// TIA Portal project "Mes_Con" (V17)

(* hardware
DEVICE "S7-1500/ET200MP station_1"  S7-1500 station
   slot 0: "Rail_0"  Rack  6ES7 590-1***0-0AA0
   slot 1: "PLC_1"  CPU 1515-2 PN  6ES7 515-2AM02-0AB0  V2.9
      slot 3: "CPU display_1"  6ES7591-1BA00-0AA0
      slot 32768: "PROFINET interface_1"  X1
         slot 32769: "Port_1"  X1 P1
         slot 32770: "Port_2"  X1 P2
      slot 33024: "PROFINET interface_2"  X2
         slot 33025: "Port_1"  X2 P1
      slot 34817: "Virtual CP interface port_1"  Virtual CP interface port  Virtual CP interface port
DEVICE "HMI_1"  KTP900 Basic PN
   slot 0: "HMI_1"  KTP900 Basic PN  6AV2 123-2JB03-0AX0  17.0.0.0
   slot 1: "HMI_RT_1"  KTP900 Basic PN  6AV2 123-2JB03-0AX0  17.0.0.0
   slot 5: "HMI_1.IE_CP_1"  PROFINET Interface  17.0.0.0
      slot 1: "PROFINET Interface_1"  PROFINET Interface
         slot 1: "Port_1"  Port
*)

// ===== PLC "PLC_1"  CPU 1515-2 PN =====

VAR_GLOBAL   // PLC tag table "Default tag table"
   "Clock_Byte" AT %MB0 : Byte;
   "Clock_10Hz" AT %M0.0 : Bool;
   "Clock_5Hz" AT %M0.1 : Bool;
   "Clock_2.5Hz" AT %M0.2 : Bool;
   "Clock_2Hz" AT %M0.3 : Bool;
   "Clock_1.25Hz" AT %M0.4 : Bool;
   "Clock_1Hz" AT %M0.5 : Bool;
   "Clock_0.625Hz" AT %M0.6 : Bool;
   "Clock_0.5Hz" AT %M0.7 : Bool;
   "System_Byte" AT %MB1 : Byte;
   "FirstScan" AT %M1.0 : Bool;
   "DiagStatusUpdate" AT %M1.1 : Bool;
   "AlwaysTRUE" AT %M1.2 : Bool;
   "AlwaysFALSE" AT %M1.3 : Bool;
   "PUMP-1_Running" AT %I10.0 : Bool;
   "PUMP-1_Thermic" AT %I10.1 : Bool;
   "PUMP-1_Loc" AT %I10.2 : Bool;
   "PUMP-2_Running" AT %I10.3 : Bool;
   "PUMP-2_Thermic" AT %I10.4 : Bool;
   "PUMP-2_Loc" AT %I10.5 : Bool;
   "PUMP-3_Running" AT %I10.6 : Bool;
   "PUMP-3_Thermic" AT %I10.7 : Bool;
   "PUMP-3_Loc" AT %I11.0 : Bool;
   "PUMP-4_Running" AT %I11.1 : Bool;
   "PUMP-4_Thermic" AT %I11.2 : Bool;
   "PUMP-4_Loc" AT %I11.3 : Bool;
   "Valve-1_Opened" AT %I11.4 : Bool;
   "Valve-1_Closed" AT %I11.5 : Bool;
   "Valve-2_Opened" AT %I11.6 : Bool;
   "Valve-2_Closed" AT %I11.7 : Bool;
   "Valve-3_Opened" AT %I12.0 : Bool;
   "Valve-3_Closed" AT %I12.1 : Bool;
   "Valve-4_Opened" AT %I12.2 : Bool;
   "Valve-4_Closed" AT %I12.3 : Bool;
   "CValve-1_Fbk" AT %IW100 : Word;
   "CValve-2_Fbk" AT %IW102 : Word;
   "CValve-3_Fbk" AT %IW104 : Word;
   "CValve-4_Fbk" AT %IW106 : Word;
   "Pump-1_RPM" AT %IW108 : Word;
   "Pump-2_RPM" AT %IW110 : Word;
   "Pump-3_RPM" AT %IW112 : Word;
   "Pump-4_RPM" AT %IW114 : Word;
   "TT-0001" AT %IW116 : Word;
   "TT-0002" AT %IW118 : Word;
   "PT-0001" AT %IW120 : Word;
   "PT-0002" AT %IW122 : Word;
   "CValve-1_Set" AT %QW200 : Word;
   "CValve-2_Set" AT %QW202 : Word;
   "CValve-3_Set" AT %QW204 : Word;
   "CValve-4_Set" AT %QW206 : Word;
   "Pump-1_SpeedRef" AT %QW208 : Word;
   "Pump-2_SpeedRef" AT %QW210 : Word;
   "Pump-3_SpeedRef" AT %QW212 : Word;
   "Pump-4_SpeedRef" AT %QW214 : Word;
   "Pump-1_Run" AT %Q50.0 : Bool;
   "Pump-2_Run" AT %Q50.1 : Bool;
   "Pump-3_Run" AT %Q50.2 : Bool;
   "Pump-4_Run" AT %Q50.3 : Bool;
   "Valve-1_Open" AT %Q50.4 : Bool;
   "Valve-2_Open" AT %Q50.5 : Bool;
   "Valve-3_Open" AT %Q50.6 : Bool;
   "Valve-4_Open" AT %Q50.7 : Bool;
   "Pump-1_Temp" AT %IW124 : Word;
   "Pump-1_A" AT %IW126 : Word;
   "Pump-2_Temp" AT %IW128 : Word;
   "Pump-2_A" AT %IW130 : Word;
   "Pump-3_Temp" AT %IW132 : Word;
   "Pump-3_A" AT %IW134 : Word;
   "Pump-4_Temp" AT %IW136 : Word;
   "Pump-4_A" AT %IW138 : Word;
END_VAR

TYPE "Popup"
VERSION : 0.1
   STRUCT
      POPUP : Array[0..99] of Bool;
   END_STRUCT;
END_TYPE

TYPE "Valve"
VERSION : 0.1
   STRUCT
      "Mod" : Bool;   // Valf Calisma durumu 0 manuel 1 otomatik
      ManuelOpen : Bool;   // MANUEL START
      ManuelClose : Bool;   // MANUEL STOP
      AutoOpen : Bool;   // AUTO START
      AutoClose : Bool;   // AUTO STOP
      Vana_Open : Bool;   // VANA AÇ
      Vana_Close : Bool;   // VANA KAPAT
      Vana_Opened : Bool;   // VANA AÇIK
      Vana_Closed : Bool;   // VANA KAPALI
      ValveStatus : Int;
      ModStatus : Int;   // VANA STATUS
      ValveIzın : Bool;
      Alarm_Not_Opened : Bool;   // AÇILMIYOR ALRM
      Alarm_Not_Closed : Bool;   // KAPANMIYOR ALARM
      Alarm_Not_Signal : Bool;   // SİNYAL YOK ALARM
      Alarm_Two_Signal : Bool;
      TimeOut : Int;   // ALARM ÇIKIŞ ZAMANI
      Alarm : Bool;   // ALARM
      Alarm_Reset : Bool;   // ALALRM RESET
      PopupClose : Bool;
      PopupInp : Bool;
      Yedek : Bool;
      Yedek_1 : Bool;
      Yedek_2 : Bool;
      Yedek_3 : Bool;
      Yedek_4 : Bool;
      Yedek_5 : Bool;
      Yedek_6 : Bool;
      Yedek_7 : Bool;
      Yedek_8 : Bool;
      Yedek_9 : Bool;
      Yedek_10 : Bool;
      Timer_1 : Int;
      Timer_2 : Int;
      Timer_4 : Int;
      Timer_5 : Int;
      Timer_3 : Int;
      Timer_6 : Int;
      Timer_7 : Int;
      Timer_8 : Int;
      Timer_9 : Int;
   END_STRUCT;
END_TYPE

TYPE "AnalogInput"
VERSION : 0.1
   STRUCT
      Input_Value : Int;
      Input_Value_Conv : Real;
      Mid_Value : Real;
      Measurement_Range : Real;
      "Procces Value_1" : Real;
      Range_Son : Real;
      Measurement_Value_Max : Real;
      Measurement_Value_Min : Real;
      Yedek_2 : Bool;
      Yedek_1 : Bool;
      Range_Control : Bool;
      AlarmTiemOut : Int := 8;
      Timer_1 : Int := 0;
      Timer_2 : Int;
      Alarm : Bool;
      Alarm_Reset : Bool;
      Range_Error : Bool;
   END_STRUCT;
END_TYPE

TYPE "AnalogOutput"
VERSION : 0.1
   STRUCT
      Process_Value : Real;
      Process_Value_Conv : Real;
      Procces_Value_Conv_Int : Int;
      Mid_Valuer : Real;
      Input_Value : Real;
      Input_Value_Real : Real;
      Measurement_Range : Real;
      Measurement_Range_Max : Real;
      Measurement_Range_Min : Real;
      RangeControl : Bool;
      Alarm : Bool;
      Range_Alarm : Bool;
      Alarm_2 : Bool;
      AlarmTimeOut : Int;
      AlarmReset : Bool;
      Yedek : Bool;
      Yedek_1 : Bool;
      Yedek_2 : Bool;
      Yedek_3 : Bool;
      Timer_1 : Int;
      Timer_3 : Int;
      Timer_2 : Int;
   END_STRUCT;
END_TYPE

TYPE "Motor"
VERSION : 0.1
   STRUCT
      "Mod" : Bool;   // 0 = Manuel Mod , 1 = Otomatik Mod
      ManuelStart : Bool;   // HMI Motor Start Button
      ManuelStop : Bool;   // HMI Motor Stop Button
      AutoStart : Bool;   // Logic Auto Start Command
      AutoStop : Bool;   // Logic Auto Stop Command
      "Local/Remote" : Bool;   // Local or Remote Button
      Motor_Rpm : Bool;
      Ucgen_Run : Bool;
      Yildiz_Run : Bool;
      iRunning : Bool;   // Motor Running Information
      iThermic : Bool;   // Motor Thermic Information
      Motor_Izın : Bool;
      Fault : Bool;   // General Fault Information
      Reset : Bool;   // Error Reset Button
      MotorStatus : Int;   // 0=Motor Calismiyor ve Hata Yok 1 = Motor Calisiyor 2 = Motor Calismasini Engelleyen Durum 3 = Motor Arıza Var
      TimeOutAlarm : Bool;   // Motor Timeout Alarm
      ThermicAlarm : Bool;   // Motor Thermic Alarm
      ShortCircuitAlarm : Bool;   // Motor Short Circuit Alarm
      MissingPhaseAlarm : Bool;   // Motor Missing Phase Alarm
      Alarm_Genel : Bool;
      Alarm6 : Bool;
      Alarm7 : Bool;
      Alarm8 : Bool;
      Yedek1 : Bool;
      Yedek2 : Bool;
      Yedek3 : Bool;
      Yedek4 : Bool;
      Yedek5 : Bool;
      Yedek6 : Bool;
      Yedek7 : Bool;
      Timer1 : Int;
      Timer2 : Int;
      Timer3 : Int;
      Timer4 : Int;
      Timer5 : Int;
      Timer6 : Int;
   END_STRUCT;
END_TYPE

TYPE "ElValve"
VERSION : 0.1
   STRUCT
      VanaOpened : Bool;
      VanaClosed : Bool;
      VanaAlarm : Bool;
      Alarm_Not_Signal : Bool;   // SİNYAL YOK ALARM
      Alarm_Two_Signal : Bool;
      Alarm_Genel : Bool;
      Alarm_Reset : Bool;
      ElV_Status : Int;
      Yedek_1 : Bool;
      Yedek_2 : Bool;
      Yedek_3 : Bool;
      Timer_1 : Int;
      Timer_2 : Int;
      Timer_3 : Int;
      TimeOut : Int;
   END_STRUCT;
END_TYPE

TYPE "FM"
VERSION : 0.1
   STRUCT
      P_Value : Real;
      Flow_Pulse_N : Int;
      F_Pulse : Bool;
      Pulse_Kg : Real;
      Total_Value : DInt;
      Set_Value : DInt;
      Tank_Value : DInt;
      TankBosaltıldı : Bool;
      SU_Alım_Run : Bool;
      TankValue_Reset : Bool;
      Total_Value_Reset : Bool;
      Pulse_Reset : Bool;
      Yedek : Bool;
      Yedek_1 : Bool;
      Yedek_2 : Int;
      Yedek_3 : Int;
   END_STRUCT;
END_TYPE

TYPE "Gunler"
VERSION : 0.1
   STRUCT
      Pazartesi : Bool;
      Salı : Bool;
      Çarşamba : Bool;
      Perşembe : Bool;
      Cuma : Bool;
      Cumartesi : Bool;
      Pazar : Bool;
      Pazartesi_Veri : Int;
      Salı_Veri : Int;
      Çarşamba_Veri : Int;
      Perşembe_Veri : Int;
      Cuma_Veri : Int;
      Cumartesi_Veri : Int;
      Pazar_Veri : Int;
      Yedek : Bool;
      Yedek_1 : Bool;
      Yedek_2 : Bool;
      Yedek_3 : Bool;
      Yedek_4 : Bool;
      Yedek_5 : Bool;
      Yedek_6 : Bool;
      Yedek_7 : Bool;
      "Timer" : Int;
      Timer_1 : Int;
      Timer_2 : Int;
      Timer_3 : Int;
   END_STRUCT;
END_TYPE

// folder: Data

DATA_BLOCK "Sim"   // DB5
{ S7_Optimized_Access := 'TRUE' }
VERSION : 0.1
   VAR
      "SPUMP-1_Running" : Bool;
      "SPUMP-1_Thermic" : Bool;
      "SPUMP-1_Loc" : Bool;
      "SPUMP-2_Running" : Bool;
      "SPUMP-2_Thermic" : Bool;
      "SPUMP-2_Loc" : Bool;
      "SPUMP-3_Running" : Bool;
      "SPUMP-3_Thermic" : Bool;
      "SPUMP-3_Loc" : Bool;
      "SPUMP-4_Running" : Bool;
      "SPUMP-4_Thermic" : Bool;
      "SPUMP-4_Loc" : Bool;
      "SValve-1_Opened" : Bool;
      "SValve-1_Closed" : Bool;
      "SValve-2_Opened" : Bool;
      "SValve-2_Closed" : Bool;
      "SValve-3_Opened" : Bool;
      "SValve-3_Closed" : Bool;
      "SValve-4_Opened" : Bool;
      "SValve-4_Closed" : Bool;
      "SPump-1_Run" : Bool;
      "SPump-2_Run" : Bool;
      "SPump-3_Run" : Bool;
      "SPump-4_Run" : Bool;
      "SValve-1_Open" : Bool;
      "SValve-2_Open" : Bool;
      "SValve-3_Open" : Bool;
      "SValve-4_Open" : Bool;
      "SCValve-1_Fbk" : Word;
      "SCValve-2_Fbk" : Word;
      "SCValve-3_Fbk" : Word;
      "SCValve-4_Fbk" : Word;
      "SPump-1_RPM" : Word;
      "SPump-2_RPM" : Word;
      "SPump-3_RPM" : Word;
      "SPump-4_RPM" : Word;
      "SPump-1_Temp" : Word;
      "SPump-1_A" : Word;
      "SPump-2_Temp" : Word;
      "SPump-2_A" : Word;
      "SPump-3_Temp" : Word;
      "SPump-3_A" : Word;
      "SPump-4_Temp" : Word;
      "SPump-4_A" : Word;
      "STT-0001" : Word;
      "STT-0002" : Word;
      "SPT-0001" : Word;
      "SPT-0002" : Word;
      "SCValve-1_Set" : Word;
      "SCValve-2_Set" : Word;
      "SCValve-3_Set" : Word;
      "SCValve-4_Set" : Word;
      "SPump-1_SpeedRef" : Word;
      "SPump-2_SpeedRef" : Word;
      "SPump-3_SpeedRef" : Word;
      "SPump-4_SpeedRef" : Word;
      SİM_MOD : Bool;
   END_VAR
BEGIN
END_DATA_BLOCK

// folder: Data/Eqp

DATA_BLOCK "PUMP"   // DB1
{ S7_Optimized_Access := 'TRUE' }
VERSION : 0.1
   VAR
      "PUMP-1" : "Motor";
      "PUMP-2" : "Motor";
      "PUMP-3" : "Motor";
      "PUMP-4" : "Motor";
   END_VAR
BEGIN
END_DATA_BLOCK

DATA_BLOCK "VALVE-H"   // DB2
{ S7_Optimized_Access := 'TRUE' }
VERSION : 0.1
   VAR
      "VALVE-1" : "Valve";
      "VALVE-2" : "Valve";
      "VALVE-3" : "Valve";
      "VALVE-4" : "Valve";
   END_VAR
BEGIN
END_DATA_BLOCK

DATA_BLOCK "VALVE-C"   // DB3
{ S7_Optimized_Access := 'TRUE' }
VERSION : 0.1
   VAR
      "CONTROLV-1" : "AnalogOutput";
      "CONTROLV-2" : "AnalogOutput";
      "CONTROLV-3" : "AnalogOutput";
      "CONTROLV-4" : "AnalogOutput";
   END_VAR
BEGIN
END_DATA_BLOCK

DATA_BLOCK "TT-PT"   // DB4
{ S7_Optimized_Access := 'TRUE' }
VERSION : 0.1
   VAR
      "TT-0001" : "AnalogInput";
      "TT-0002" : "AnalogInput";
      "PT-0001" : "AnalogInput";
      "PT-0002" : "AnalogInput";
   END_VAR
BEGIN
END_DATA_BLOCK

// folder: Data/HMI

DATA_BLOCK "HMI"   // DB7
{ S7_Optimized_Access := 'TRUE' }
VERSION : 0.1
   VAR
      Popup : "Popup";
      "CValve-1_Set" : Int;
      "CValve-2_Set" : Int;
      "CValve-3_Set" : Int;
      "CValve-4_Set" : Int;
      "Pump-1" : Int;
      "Pump-2" : Int;
      "Pump-3" : Int;
      "Pump-4" : Int;
   END_VAR
BEGIN
END_DATA_BLOCK

// folder: Data/mes

DATA_BLOCK "Connection"   // DB6
{ S7_Optimized_Access := 'FALSE' }
VERSION : 0.1
   VAR
      "CV-1Flt" : Bool;
      "CV-2Flt" : Bool;
      "CV-3Flt" : Bool;
      "CV-4Flt" : Bool;
      "TT1-FLT" : Bool;
      "TT2-FLT" : Bool;
      "PT1-FLT" : Bool;
      "PT2-FLT" : Bool;
      "Pump-1Status" : Word;
      "Pump-2Status" : Word;
      "Pump-3Status" : Word;
      "Pump-4Status" : Word;
      "V1-Status" : Word;
      "V2-Status" : Word;
      "V3-Status" : Word;
      "V4-Status" : Word;
      "Pump1-Rpm" : Word;
      "Pump2-Rpm" : Word;
      "Pump3-Rpm" : Word;
      "Pump4-Rpm" : Word;
      "CV1-Percent" : Word;
      "CV2-Percent" : Word;
      "CV3-Percent" : Word;
      "CV4-Percent" : Word;
      "TT1-Value" : Word;
      "TT2-Value" : Word;
      "PT1-Value" : Word;
      "PT2-Value" : Word;
   END_VAR
BEGIN
END_DATA_BLOCK

DATA_BLOCK "workorder"   // DB10
{ S7_Optimized_Access := 'FALSE' }
VERSION : 0.1
   VAR
      "Work_Order-1_Active" : Bool;
      "Work_Order-2_Active" : Bool;
      "Work_Order-3_Active" : Bool;
      "Work_Order-4_Active" : Bool;
      "Work_Order-5_Active" : Bool;
      "Work_Order-6_Active" : Bool;
      "Work_Order-7_Active" : Bool;
      "Work_Order-8_Active" : Bool;
      "Work_Order-9_Active" : Bool;
      "Work_Order-10_Active" : Bool;
      "Work_Order-11_Active" : Bool;
      "Work_Order-12_Active" : Bool;
      "Work_Order-13_Active" : Bool;
      "Work_Order-14_Active" : Bool;
      "Work_Order-15_Active" : Bool;
   END_VAR
BEGIN
END_DATA_BLOCK

DATA_BLOCK "maint"   // DB100
{ S7_Optimized_Access := 'TRUE' }
VERSION : 0.1
   VAR
      "Pump-1_Sim" : Bool;
      "Pump-1_Running" : Bool;
      "Pump-1_Loc" : Bool;
      "Pump-1_PhaseAlarm" : Bool;
      "Pump-1_ThermicAlarm" : Bool;
      "Pump-1_TimeOutAlarm" : Bool;
      "Pump-1_ShortCircuit" : Bool;
      "Pump-2_Sim" : Bool;
      "Pump-2_Running" : Bool;
      "Pump-2_Loc" : Bool;
      "Pump-2_PhaseAlarm" : Bool;
      "Pump-2_ThermicAlarm" : Bool;
      "Pump-2_TimeOutAlarm" : Bool;
      "Pump-2_ShortCircuit" : Bool;
      "Pump-3_Sim" : Bool;
      "Pump-3_Running" : Bool;
      "Pump-3_Loc" : Bool;
      "Pump-3_PhaseAlarm" : Bool;
      "Pump-3_ThermicAlarm" : Bool;
      "Pump-3_TimeOutAlarm" : Bool;
      "Pump-3_ShortCircuit" : Bool;
      "Pump-4_Sim" : Bool;
      "Pump-4_Running" : Bool;
      "Pump-4_Loc" : Bool;
      "Pump-4_PhaseAlarm" : Bool;
      "Pump-4_ThermicAlarm" : Bool;
      "Pump-4_TimeOutAlarm" : Bool;
      "Pump-4_ShortCircuit" : Bool;
      "Valve-1_Sim" : Bool;
      "Valve-1_NotOpened" : Bool;
      "Valve-1_NotClosed" : Bool;
      "Valve-1_NotSignal" : Bool;
      "Valve-1_TwoSignal" : Bool;
      "Valve-2_Sim" : Bool;
      "Valve-2_NotOpened" : Bool;
      "Valve-2_NotClosed" : Bool;
      "Valve-2_NotSignal" : Bool;
      "Valve-2_TwoSignal" : Bool;
      "Valve-3_Sim" : Bool;
      "Valve-3_NotOpened" : Bool;
      "Valve-3_NotClosed" : Bool;
      "Valve-3_NotSignal" : Bool;
      "Valve-3_TwoSignal" : Bool;
      "Valve-4_Sim" : Bool;
      "Valve-4_NotOpened" : Bool;
      "Valve-4_NotClosed" : Bool;
      "Valve-4_NotSignal" : Bool;
      "Valve-4_TwoSignal" : Bool;
      "Pump-1_A" : Word;
      "Pump-1_Temp" : Word;
      "Pump-2_A" : Word;
      "Pump-2_Temp" : Word;
      "Pump-3_A" : Word;
      "Pump-3_Temp" : Word;
      "Pump-4_A" : Word;
      "Pump-4_Temp" : Word;
      "TT-0001" : Word;
      "TT-0002" : Word;
      "PT-0001" : Word;
      "PT-0002" : Word;
      "CValve-1_FBK" : Word;
      "CValve-2_FBK" : Word;
      "CValve-3_FBK" : Word;
      "CValve-4_FBK" : Word;
   END_VAR
BEGIN
END_DATA_BLOCK

// folder: (top level)

FUNCTION "Equipment" : Void   // FC2, LAD
{ S7_Optimized_Access := 'TRUE' }
VERSION : 0.1
BEGIN

REGION Network 1: PUMP-1
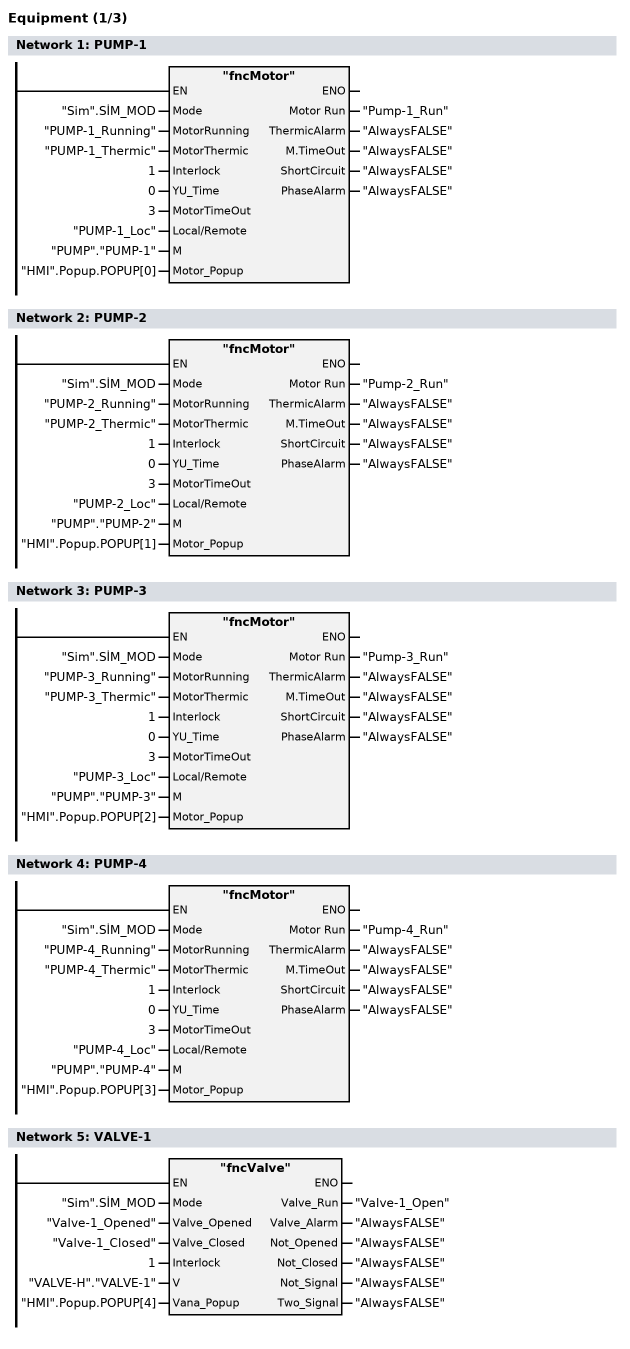
   RUNG wire#powerrail
      "fncMotor"(Mode := "Sim".SİM_MOD, MotorRunning := "PUMP-1_Running", MotorThermic := "PUMP-1_Thermic", Interlock := 1, YU_Time := 0, MotorTimeOut := 3, "Local/Remote" := "PUMP-1_Loc", "M" := "PUMP"."PUMP-1", Motor_Popup := "HMI".Popup.POPUP[0], "Motor Run" => "Pump-1_Run", ThermicAlarm => "AlwaysFALSE", "M.TimeOut" => "AlwaysFALSE", ShortCircuit => "AlwaysFALSE", PhaseAlarm => "AlwaysFALSE")
   END_RUNG
   // the same network as SCL:
   "fncMotor"(Mode := "Sim".SİM_MOD,
              MotorRunning := "PUMP-1_Running",
              MotorThermic := "PUMP-1_Thermic",
              Interlock := 1,
              YU_Time := 0,
              MotorTimeOut := 3,
              "Local/Remote" := "PUMP-1_Loc",
              "M" := "PUMP"."PUMP-1",
              Motor_Popup := "HMI".Popup.POPUP[0],
              "Motor Run" => "Pump-1_Run",
              ThermicAlarm => "AlwaysFALSE",
              "M.TimeOut" => "AlwaysFALSE",
              ShortCircuit => "AlwaysFALSE",
              PhaseAlarm => "AlwaysFALSE");
END_REGION

REGION Network 2: PUMP-2
   RUNG wire#powerrail
      "fncMotor"(Mode := "Sim".SİM_MOD, MotorRunning := "PUMP-2_Running", MotorThermic := "PUMP-2_Thermic", Interlock := 1, YU_Time := 0, MotorTimeOut := 3, "Local/Remote" := "PUMP-2_Loc", "M" := "PUMP"."PUMP-2", Motor_Popup := "HMI".Popup.POPUP[1], "Motor Run" => "Pump-2_Run", ThermicAlarm => "AlwaysFALSE", "M.TimeOut" => "AlwaysFALSE", ShortCircuit => "AlwaysFALSE", PhaseAlarm => "AlwaysFALSE")
   END_RUNG
   // the same network as SCL:
   "fncMotor"(Mode := "Sim".SİM_MOD,
              MotorRunning := "PUMP-2_Running",
              MotorThermic := "PUMP-2_Thermic",
              Interlock := 1,
              YU_Time := 0,
              MotorTimeOut := 3,
              "Local/Remote" := "PUMP-2_Loc",
              "M" := "PUMP"."PUMP-2",
              Motor_Popup := "HMI".Popup.POPUP[1],
              "Motor Run" => "Pump-2_Run",
              ThermicAlarm => "AlwaysFALSE",
              "M.TimeOut" => "AlwaysFALSE",
              ShortCircuit => "AlwaysFALSE",
              PhaseAlarm => "AlwaysFALSE");
END_REGION

REGION Network 3: PUMP-3
   RUNG wire#powerrail
      "fncMotor"(Mode := "Sim".SİM_MOD, MotorRunning := "PUMP-3_Running", MotorThermic := "PUMP-3_Thermic", Interlock := 1, YU_Time := 0, MotorTimeOut := 3, "Local/Remote" := "PUMP-3_Loc", "M" := "PUMP"."PUMP-3", Motor_Popup := "HMI".Popup.POPUP[2], "Motor Run" => "Pump-3_Run", ThermicAlarm => "AlwaysFALSE", "M.TimeOut" => "AlwaysFALSE", ShortCircuit => "AlwaysFALSE", PhaseAlarm => "AlwaysFALSE")
   END_RUNG
   // the same network as SCL:
   "fncMotor"(Mode := "Sim".SİM_MOD,
              MotorRunning := "PUMP-3_Running",
              MotorThermic := "PUMP-3_Thermic",
              Interlock := 1,
              YU_Time := 0,
              MotorTimeOut := 3,
              "Local/Remote" := "PUMP-3_Loc",
              "M" := "PUMP"."PUMP-3",
              Motor_Popup := "HMI".Popup.POPUP[2],
              "Motor Run" => "Pump-3_Run",
              ThermicAlarm => "AlwaysFALSE",
              "M.TimeOut" => "AlwaysFALSE",
              ShortCircuit => "AlwaysFALSE",
              PhaseAlarm => "AlwaysFALSE");
END_REGION

REGION Network 4: PUMP-4
   RUNG wire#powerrail
      "fncMotor"(Mode := "Sim".SİM_MOD, MotorRunning := "PUMP-4_Running", MotorThermic := "PUMP-4_Thermic", Interlock := 1, YU_Time := 0, MotorTimeOut := 3, "Local/Remote" := "PUMP-4_Loc", "M" := "PUMP"."PUMP-4", Motor_Popup := "HMI".Popup.POPUP[3], "Motor Run" => "Pump-4_Run", ThermicAlarm => "AlwaysFALSE", "M.TimeOut" => "AlwaysFALSE", ShortCircuit => "AlwaysFALSE", PhaseAlarm => "AlwaysFALSE")
   END_RUNG
   // the same network as SCL:
   "fncMotor"(Mode := "Sim".SİM_MOD,
              MotorRunning := "PUMP-4_Running",
              MotorThermic := "PUMP-4_Thermic",
              Interlock := 1,
              YU_Time := 0,
              MotorTimeOut := 3,
              "Local/Remote" := "PUMP-4_Loc",
              "M" := "PUMP"."PUMP-4",
              Motor_Popup := "HMI".Popup.POPUP[3],
              "Motor Run" => "Pump-4_Run",
              ThermicAlarm => "AlwaysFALSE",
              "M.TimeOut" => "AlwaysFALSE",
              ShortCircuit => "AlwaysFALSE",
              PhaseAlarm => "AlwaysFALSE");
END_REGION

REGION Network 5: VALVE-1
   RUNG wire#powerrail
      "fncValve"(Mode := "Sim".SİM_MOD, Valve_Opened := "Valve-1_Opened", Valve_Closed := "Valve-1_Closed", Interlock := 1, V := "VALVE-H"."VALVE-1", Vana_Popup := "HMI".Popup.POPUP[4], Valve_Run => "Valve-1_Open", Valve_Alarm => "AlwaysFALSE", Not_Opened => "AlwaysFALSE", Not_Closed => "AlwaysFALSE", Not_Signal => "AlwaysFALSE", Two_Signal => "AlwaysFALSE")
   END_RUNG
   // the same network as SCL:
   "fncValve"(Mode := "Sim".SİM_MOD,
              Valve_Opened := "Valve-1_Opened",
              Valve_Closed := "Valve-1_Closed",
              Interlock := 1,
              V := "VALVE-H"."VALVE-1",
              Vana_Popup := "HMI".Popup.POPUP[4],
              Valve_Run => "Valve-1_Open",
              Valve_Alarm => "AlwaysFALSE",
              Not_Opened => "AlwaysFALSE",
              Not_Closed => "AlwaysFALSE",
              Not_Signal => "AlwaysFALSE",
              Two_Signal => "AlwaysFALSE");
END_REGION

REGION Network 6: VALVE-2
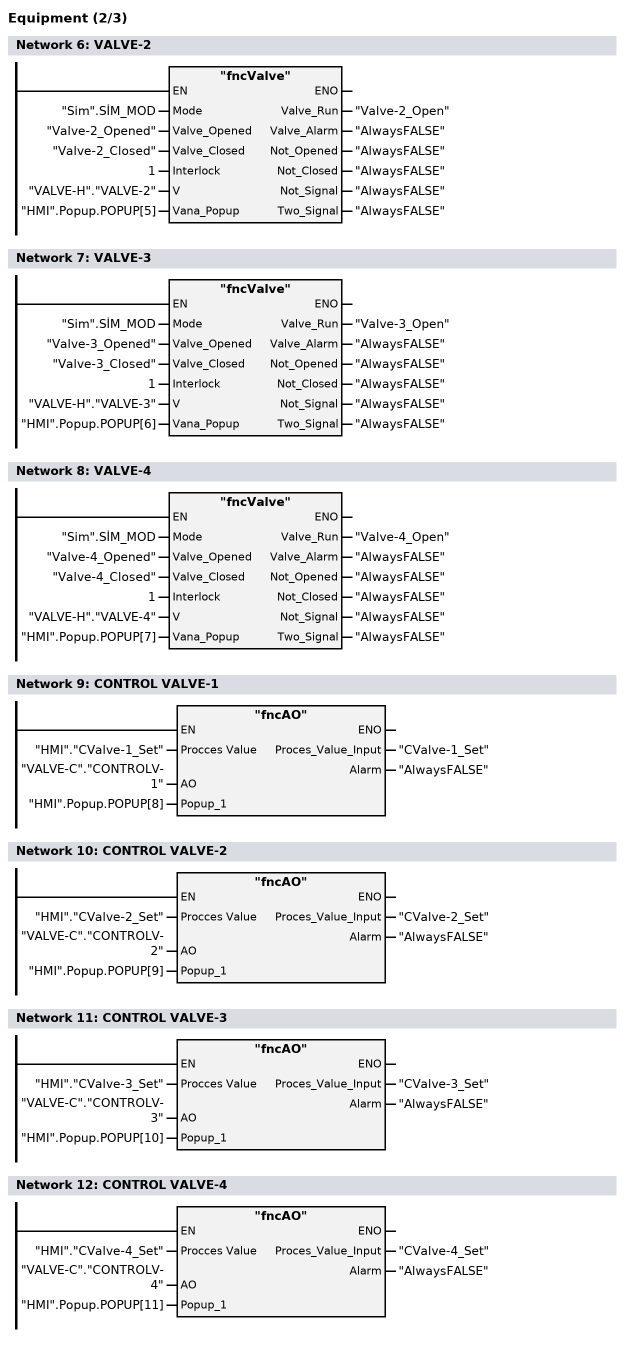
   RUNG wire#powerrail
      "fncValve"(Mode := "Sim".SİM_MOD, Valve_Opened := "Valve-2_Opened", Valve_Closed := "Valve-2_Closed", Interlock := 1, V := "VALVE-H"."VALVE-2", Vana_Popup := "HMI".Popup.POPUP[5], Valve_Run => "Valve-2_Open", Valve_Alarm => "AlwaysFALSE", Not_Opened => "AlwaysFALSE", Not_Closed => "AlwaysFALSE", Not_Signal => "AlwaysFALSE", Two_Signal => "AlwaysFALSE")
   END_RUNG
   // the same network as SCL:
   "fncValve"(Mode := "Sim".SİM_MOD,
              Valve_Opened := "Valve-2_Opened",
              Valve_Closed := "Valve-2_Closed",
              Interlock := 1,
              V := "VALVE-H"."VALVE-2",
              Vana_Popup := "HMI".Popup.POPUP[5],
              Valve_Run => "Valve-2_Open",
              Valve_Alarm => "AlwaysFALSE",
              Not_Opened => "AlwaysFALSE",
              Not_Closed => "AlwaysFALSE",
              Not_Signal => "AlwaysFALSE",
              Two_Signal => "AlwaysFALSE");
END_REGION

REGION Network 7: VALVE-3
   RUNG wire#powerrail
      "fncValve"(Mode := "Sim".SİM_MOD, Valve_Opened := "Valve-3_Opened", Valve_Closed := "Valve-3_Closed", Interlock := 1, V := "VALVE-H"."VALVE-3", Vana_Popup := "HMI".Popup.POPUP[6], Valve_Run => "Valve-3_Open", Valve_Alarm => "AlwaysFALSE", Not_Opened => "AlwaysFALSE", Not_Closed => "AlwaysFALSE", Not_Signal => "AlwaysFALSE", Two_Signal => "AlwaysFALSE")
   END_RUNG
   // the same network as SCL:
   "fncValve"(Mode := "Sim".SİM_MOD,
              Valve_Opened := "Valve-3_Opened",
              Valve_Closed := "Valve-3_Closed",
              Interlock := 1,
              V := "VALVE-H"."VALVE-3",
              Vana_Popup := "HMI".Popup.POPUP[6],
              Valve_Run => "Valve-3_Open",
              Valve_Alarm => "AlwaysFALSE",
              Not_Opened => "AlwaysFALSE",
              Not_Closed => "AlwaysFALSE",
              Not_Signal => "AlwaysFALSE",
              Two_Signal => "AlwaysFALSE");
END_REGION

REGION Network 8: VALVE-4
   RUNG wire#powerrail
      "fncValve"(Mode := "Sim".SİM_MOD, Valve_Opened := "Valve-4_Opened", Valve_Closed := "Valve-4_Closed", Interlock := 1, V := "VALVE-H"."VALVE-4", Vana_Popup := "HMI".Popup.POPUP[7], Valve_Run => "Valve-4_Open", Valve_Alarm => "AlwaysFALSE", Not_Opened => "AlwaysFALSE", Not_Closed => "AlwaysFALSE", Not_Signal => "AlwaysFALSE", Two_Signal => "AlwaysFALSE")
   END_RUNG
   // the same network as SCL:
   "fncValve"(Mode := "Sim".SİM_MOD,
              Valve_Opened := "Valve-4_Opened",
              Valve_Closed := "Valve-4_Closed",
              Interlock := 1,
              V := "VALVE-H"."VALVE-4",
              Vana_Popup := "HMI".Popup.POPUP[7],
              Valve_Run => "Valve-4_Open",
              Valve_Alarm => "AlwaysFALSE",
              Not_Opened => "AlwaysFALSE",
              Not_Closed => "AlwaysFALSE",
              Not_Signal => "AlwaysFALSE",
              Two_Signal => "AlwaysFALSE");
END_REGION

REGION Network 9: CONTROL VALVE-1
   RUNG wire#powerrail
      "fncAO"("Procces Value" := "HMI"."CValve-1_Set", AO := "VALVE-C"."CONTROLV-1", Popup_1 := "HMI".Popup.POPUP[8], Proces_Value_Input => "CValve-1_Set", Alarm => "AlwaysFALSE")
   END_RUNG
   // the same network as SCL:
   "fncAO"("Procces Value" := "HMI"."CValve-1_Set",
           AO := "VALVE-C"."CONTROLV-1",
           Popup_1 := "HMI".Popup.POPUP[8],
           Proces_Value_Input => "CValve-1_Set",
           Alarm => "AlwaysFALSE");
END_REGION

REGION Network 10: CONTROL VALVE-2
   RUNG wire#powerrail
      "fncAO"("Procces Value" := "HMI"."CValve-2_Set", AO := "VALVE-C"."CONTROLV-2", Popup_1 := "HMI".Popup.POPUP[9], Proces_Value_Input => "CValve-2_Set", Alarm => "AlwaysFALSE")
   END_RUNG
   // the same network as SCL:
   "fncAO"("Procces Value" := "HMI"."CValve-2_Set",
           AO := "VALVE-C"."CONTROLV-2",
           Popup_1 := "HMI".Popup.POPUP[9],
           Proces_Value_Input => "CValve-2_Set",
           Alarm => "AlwaysFALSE");
END_REGION

REGION Network 11: CONTROL VALVE-3
   RUNG wire#powerrail
      "fncAO"("Procces Value" := "HMI"."CValve-3_Set", AO := "VALVE-C"."CONTROLV-3", Popup_1 := "HMI".Popup.POPUP[10], Proces_Value_Input => "CValve-3_Set", Alarm => "AlwaysFALSE")
   END_RUNG
   // the same network as SCL:
   "fncAO"("Procces Value" := "HMI"."CValve-3_Set",
           AO := "VALVE-C"."CONTROLV-3",
           Popup_1 := "HMI".Popup.POPUP[10],
           Proces_Value_Input => "CValve-3_Set",
           Alarm => "AlwaysFALSE");
END_REGION

REGION Network 12: CONTROL VALVE-4
   RUNG wire#powerrail
      "fncAO"("Procces Value" := "HMI"."CValve-4_Set", AO := "VALVE-C"."CONTROLV-4", Popup_1 := "HMI".Popup.POPUP[11], Proces_Value_Input => "CValve-4_Set", Alarm => "AlwaysFALSE")
   END_RUNG
   // the same network as SCL:
   "fncAO"("Procces Value" := "HMI"."CValve-4_Set",
           AO := "VALVE-C"."CONTROLV-4",
           Popup_1 := "HMI".Popup.POPUP[11],
           Proces_Value_Input => "CValve-4_Set",
           Alarm => "AlwaysFALSE");
END_REGION

REGION Network 13: TT-0001
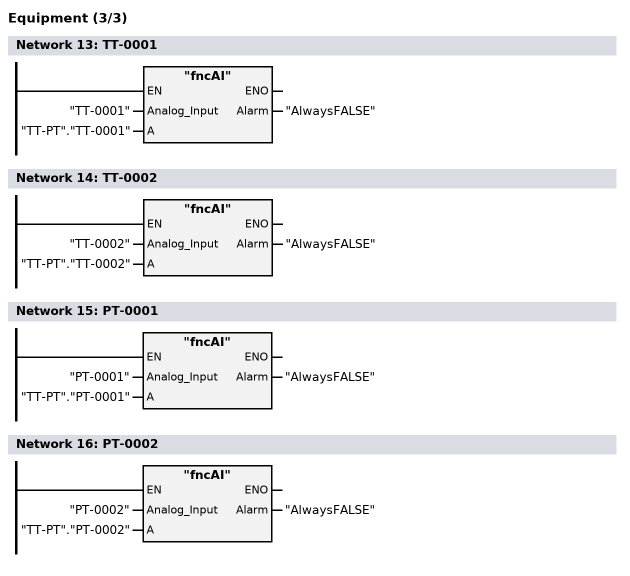
   RUNG wire#powerrail
      "fncAI"(Analog_Input := "TT-0001", "A" := "TT-PT"."TT-0001", Alarm => "AlwaysFALSE")
   END_RUNG
   // the same network as SCL:
   "fncAI"(Analog_Input := "TT-0001", "A" := "TT-PT"."TT-0001", Alarm => "AlwaysFALSE");
END_REGION

REGION Network 14: TT-0002
   RUNG wire#powerrail
      "fncAI"(Analog_Input := "TT-0002", "A" := "TT-PT"."TT-0002", Alarm => "AlwaysFALSE")
   END_RUNG
   // the same network as SCL:
   "fncAI"(Analog_Input := "TT-0002", "A" := "TT-PT"."TT-0002", Alarm => "AlwaysFALSE");
END_REGION

REGION Network 15: PT-0001
   RUNG wire#powerrail
      "fncAI"(Analog_Input := "PT-0001", "A" := "TT-PT"."PT-0001", Alarm => "AlwaysFALSE")
   END_RUNG
   // the same network as SCL:
   "fncAI"(Analog_Input := "PT-0001", "A" := "TT-PT"."PT-0001", Alarm => "AlwaysFALSE");
END_REGION

REGION Network 16: PT-0002
   RUNG wire#powerrail
      "fncAI"(Analog_Input := "PT-0002", "A" := "TT-PT"."PT-0002", Alarm => "AlwaysFALSE")
   END_RUNG
   // the same network as SCL:
   "fncAI"(Analog_Input := "PT-0002", "A" := "TT-PT"."PT-0002", Alarm => "AlwaysFALSE");
END_REGION
END_FUNCTION

FUNCTION "Simfnc" : Void   // FC19, LAD
{ S7_Optimized_Access := 'TRUE' }
VERSION : 0.1
BEGIN

REGION Network 1: PUMP-1
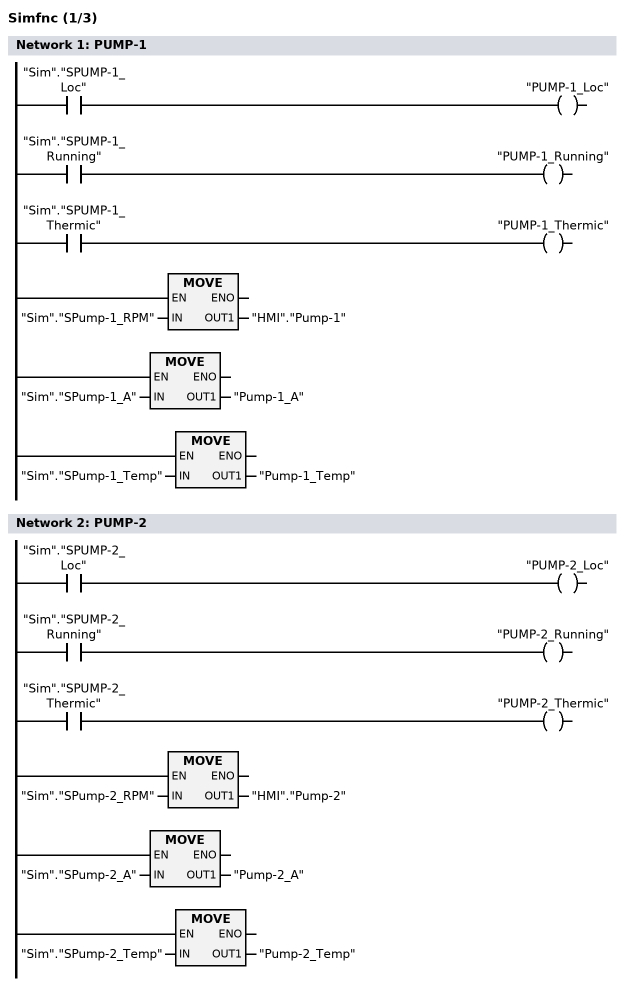
   RUNG wire#powerrail
      Contact( "Sim"."SPUMP-1_Loc" )
      Coil( "PUMP-1_Loc" )
   END_RUNG
   RUNG wire#powerrail
      Contact( "Sim"."SPUMP-1_Running" )
      Coil( "PUMP-1_Running" )
   END_RUNG
   RUNG wire#powerrail
      Contact( "Sim"."SPUMP-1_Thermic" )
      Coil( "PUMP-1_Thermic" )
   END_RUNG
   RUNG wire#powerrail
      Move(in := "Sim"."SPump-1_RPM", out1 => "HMI"."Pump-1")
   END_RUNG
   RUNG wire#powerrail
      Move(in := "Sim"."SPump-1_A", out1 => "Pump-1_A")
   END_RUNG
   RUNG wire#powerrail
      Move(in := "Sim"."SPump-1_Temp", out1 => "Pump-1_Temp")
   END_RUNG
   // the same network as SCL:
   "PUMP-1_Loc" := "Sim"."SPUMP-1_Loc";
   "PUMP-1_Running" := "Sim"."SPUMP-1_Running";
   "PUMP-1_Thermic" := "Sim"."SPUMP-1_Thermic";
   "HMI"."Pump-1" := "Sim"."SPump-1_RPM";
   "Pump-1_A" := "Sim"."SPump-1_A";
   "Pump-1_Temp" := "Sim"."SPump-1_Temp";
END_REGION

REGION Network 2: PUMP-2
   RUNG wire#powerrail
      Contact( "Sim"."SPUMP-2_Loc" )
      Coil( "PUMP-2_Loc" )
   END_RUNG
   RUNG wire#powerrail
      Contact( "Sim"."SPUMP-2_Running" )
      Coil( "PUMP-2_Running" )
   END_RUNG
   RUNG wire#powerrail
      Contact( "Sim"."SPUMP-2_Thermic" )
      Coil( "PUMP-2_Thermic" )
   END_RUNG
   RUNG wire#powerrail
      Move(in := "Sim"."SPump-2_RPM", out1 => "HMI"."Pump-2")
   END_RUNG
   RUNG wire#powerrail
      Move(in := "Sim"."SPump-2_A", out1 => "Pump-2_A")
   END_RUNG
   RUNG wire#powerrail
      Move(in := "Sim"."SPump-2_Temp", out1 => "Pump-2_Temp")
   END_RUNG
   // the same network as SCL:
   "PUMP-2_Loc" := "Sim"."SPUMP-2_Loc";
   "PUMP-2_Running" := "Sim"."SPUMP-2_Running";
   "PUMP-2_Thermic" := "Sim"."SPUMP-2_Thermic";
   "HMI"."Pump-2" := "Sim"."SPump-2_RPM";
   "Pump-2_A" := "Sim"."SPump-2_A";
   "Pump-2_Temp" := "Sim"."SPump-2_Temp";
END_REGION

REGION Network 3: PUMP-3
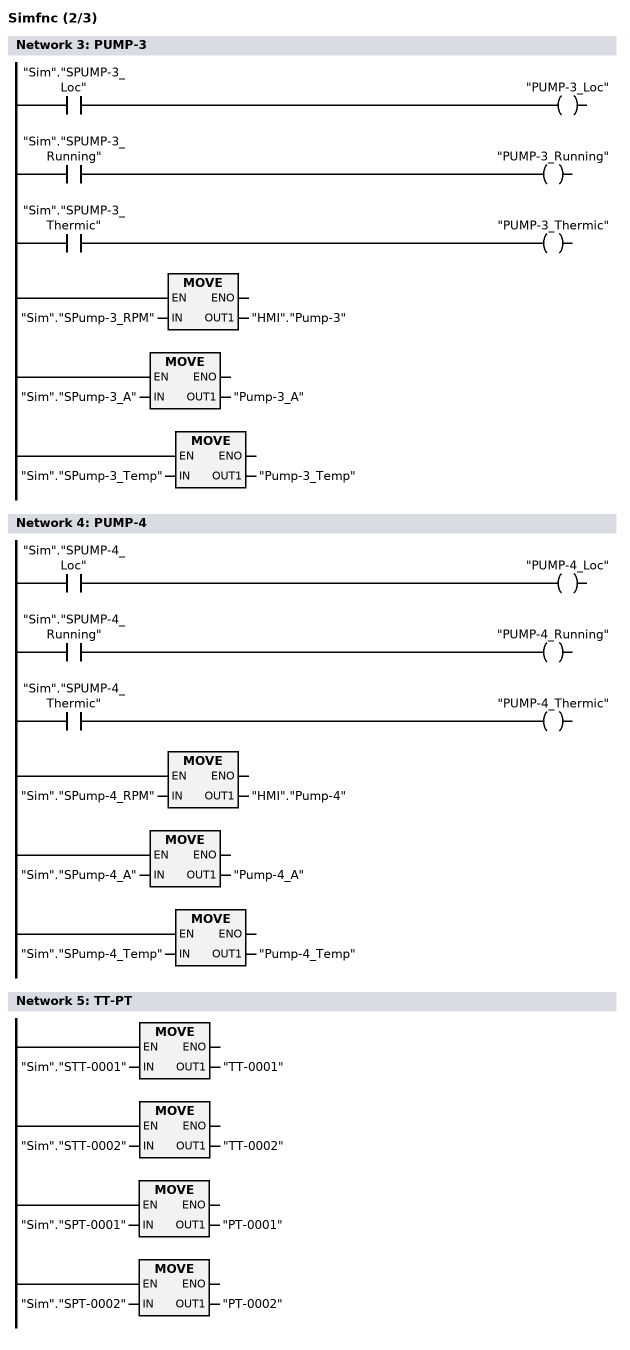
   RUNG wire#powerrail
      Contact( "Sim"."SPUMP-3_Loc" )
      Coil( "PUMP-3_Loc" )
   END_RUNG
   RUNG wire#powerrail
      Contact( "Sim"."SPUMP-3_Running" )
      Coil( "PUMP-3_Running" )
   END_RUNG
   RUNG wire#powerrail
      Contact( "Sim"."SPUMP-3_Thermic" )
      Coil( "PUMP-3_Thermic" )
   END_RUNG
   RUNG wire#powerrail
      Move(in := "Sim"."SPump-3_RPM", out1 => "HMI"."Pump-3")
   END_RUNG
   RUNG wire#powerrail
      Move(in := "Sim"."SPump-3_A", out1 => "Pump-3_A")
   END_RUNG
   RUNG wire#powerrail
      Move(in := "Sim"."SPump-3_Temp", out1 => "Pump-3_Temp")
   END_RUNG
   // the same network as SCL:
   "PUMP-3_Loc" := "Sim"."SPUMP-3_Loc";
   "PUMP-3_Running" := "Sim"."SPUMP-3_Running";
   "PUMP-3_Thermic" := "Sim"."SPUMP-3_Thermic";
   "HMI"."Pump-3" := "Sim"."SPump-3_RPM";
   "Pump-3_A" := "Sim"."SPump-3_A";
   "Pump-3_Temp" := "Sim"."SPump-3_Temp";
END_REGION

REGION Network 4: PUMP-4
   RUNG wire#powerrail
      Contact( "Sim"."SPUMP-4_Loc" )
      Coil( "PUMP-4_Loc" )
   END_RUNG
   RUNG wire#powerrail
      Contact( "Sim"."SPUMP-4_Running" )
      Coil( "PUMP-4_Running" )
   END_RUNG
   RUNG wire#powerrail
      Contact( "Sim"."SPUMP-4_Thermic" )
      Coil( "PUMP-4_Thermic" )
   END_RUNG
   RUNG wire#powerrail
      Move(in := "Sim"."SPump-4_RPM", out1 => "HMI"."Pump-4")
   END_RUNG
   RUNG wire#powerrail
      Move(in := "Sim"."SPump-4_A", out1 => "Pump-4_A")
   END_RUNG
   RUNG wire#powerrail
      Move(in := "Sim"."SPump-4_Temp", out1 => "Pump-4_Temp")
   END_RUNG
   // the same network as SCL:
   "PUMP-4_Loc" := "Sim"."SPUMP-4_Loc";
   "PUMP-4_Running" := "Sim"."SPUMP-4_Running";
   "PUMP-4_Thermic" := "Sim"."SPUMP-4_Thermic";
   "HMI"."Pump-4" := "Sim"."SPump-4_RPM";
   "Pump-4_A" := "Sim"."SPump-4_A";
   "Pump-4_Temp" := "Sim"."SPump-4_Temp";
END_REGION

REGION Network 5: TT-PT
   RUNG wire#powerrail
      Move(in := "Sim"."STT-0001", out1 => "TT-0001")
   END_RUNG
   RUNG wire#powerrail
      Move(in := "Sim"."STT-0002", out1 => "TT-0002")
   END_RUNG
   RUNG wire#powerrail
      Move(in := "Sim"."SPT-0001", out1 => "PT-0001")
   END_RUNG
   RUNG wire#powerrail
      Move(in := "Sim"."SPT-0002", out1 => "PT-0002")
   END_RUNG
   // the same network as SCL:
   "TT-0001" := "Sim"."STT-0001";
   "TT-0002" := "Sim"."STT-0002";
   "PT-0001" := "Sim"."SPT-0001";
   "PT-0002" := "Sim"."SPT-0002";
END_REGION

REGION Network 6: CVALVE FBK
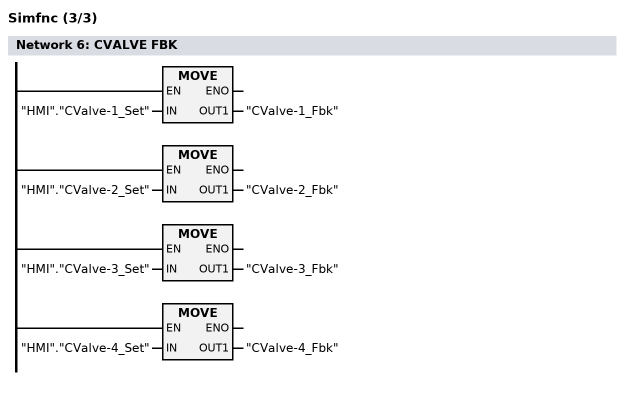
   RUNG wire#powerrail
      Move(in := "HMI"."CValve-1_Set", out1 => "CValve-1_Fbk")
   END_RUNG
   RUNG wire#powerrail
      Move(in := "HMI"."CValve-2_Set", out1 => "CValve-2_Fbk")
   END_RUNG
   RUNG wire#powerrail
      Move(in := "HMI"."CValve-3_Set", out1 => "CValve-3_Fbk")
   END_RUNG
   RUNG wire#powerrail
      Move(in := "HMI"."CValve-4_Set", out1 => "CValve-4_Fbk")
   END_RUNG
   // the same network as SCL:
   "CValve-1_Fbk" := "HMI"."CValve-1_Set";
   "CValve-2_Fbk" := "HMI"."CValve-2_Set";
   "CValve-3_Fbk" := "HMI"."CValve-3_Set";
   "CValve-4_Fbk" := "HMI"."CValve-4_Set";
END_REGION
END_FUNCTION

ORGANIZATION_BLOCK "Main"   // OB1, LAD, ProgramCycle
TITLE = "Main Program Sweep (Cycle)"
{ S7_Optimized_Access := 'TRUE' }
VERSION : 0.1
   VAR_INPUT
      Initial_Call : Bool;   // Initial call of this OB
      Remanence : Bool;   // =True, if remanent data are available
   END_VAR
BEGIN

REGION Network 1
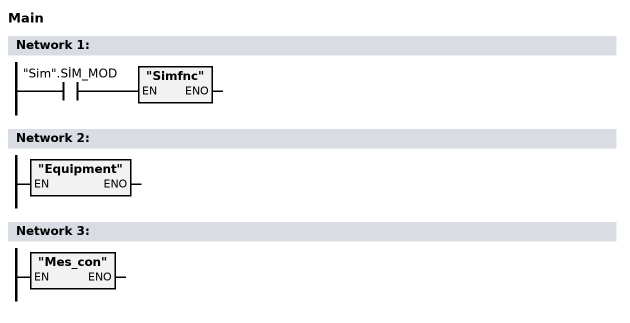
   RUNG wire#powerrail
      Contact( "Sim".SİM_MOD )
      "Simfnc"()
   END_RUNG
   // the same network as SCL:
   IF "Sim".SİM_MOD THEN "Simfnc"(); END_IF;
END_REGION

REGION Network 2
   RUNG wire#powerrail
      "Equipment"()
   END_RUNG
   // the same network as SCL:
   "Equipment"();
END_REGION

REGION Network 3
   RUNG wire#powerrail
      "Mes_con"()
   END_RUNG
   // the same network as SCL:
   "Mes_con"();
END_REGION
END_ORGANIZATION_BLOCK

// folder: Data/mes

FUNCTION "Mes_con" : Void   // FC4, LAD
{ S7_Optimized_Access := 'TRUE' }
VERSION : 0.1
BEGIN

REGION Network 1: PUMP